REGION Network 18: I21.1 - Tank Group Pressure HIHI (PS-436)
   // True = OK, False = HIHI
   RUNG wire#powerrail
      I_Contact( "RIO2 Tanks Pressure Switch Hi Hi" )
      Coil( "20_TANKS_IP_DATA".RIO_02.FIRST_TANK.TANKS_PRESS_HIHI )
   END_RUNG
   // the same network as SCL:
   "20_TANKS_IP_DATA".RIO_02.FIRST_TANK.TANKS_PRESS_HIHI := NOT "RIO2 Tanks Pressure Switch Hi Hi";
END_REGION

REGION Network 19: I21.2 - Tank Level HIHI - (LS-425) - Second Tank
   // True = OK, False = HIHI
   RUNG wire#powerrail
      I_Contact( "Tank 2S BWT Level High High Switch" )
      Coil( "20_TANKS_IP_DATA".RIO_02.SECOND_TANK.BWT_LEVEL_HIHI )
   END_RUNG
   // the same network as SCL:
   "20_TANKS_IP_DATA".RIO_02.SECOND_TANK.BWT_LEVEL_HIHI := NOT "Tank 2S BWT Level High High Switch";
END_REGION

REGION Network 20: I21.3 - Spare Input
   // True = N/A, False = N/A
   RUNG wire#powerrail
      Contact( "RIO2_SPR_DI_21_3" )
      Coil( "20_TANKS_IP_DATA".RIO_02.FIRST_TANK.TANK_GROUP_SPARE_DI_3 )
   END_RUNG
   // the same network as SCL:
   "20_TANKS_IP_DATA".RIO_02.FIRST_TANK.TANK_GROUP_SPARE_DI_3 := "RIO2_SPR_DI_21_3";
END_REGION

REGION Network 21: I21.4 - Spare Input
   // True = N/A, False = N/A
   RUNG wire#powerrail
      Contact( "RIO2_SPR_DI_21_4" )
      Coil( "20_TANKS_IP_DATA".RIO_02.FIRST_TANK.TANK_GROUP_SPARE_DI_4 )
   END_RUNG
   // the same network as SCL:
   "20_TANKS_IP_DATA".RIO_02.FIRST_TANK.TANK_GROUP_SPARE_DI_4 := "RIO2_SPR_DI_21_4";
END_REGION

REGION Network 22: I21.5 - Spare Input
   // True = N/A, False = N/A
   RUNG wire#powerrail
      Contact( "RIO2_SPR_DI_21_5" )
      Coil( "20_TANKS_IP_DATA".RIO_02.FIRST_TANK.TANK_GROUP_SPARE_DI_5 )
   END_RUNG
   // the same network as SCL:
   "20_TANKS_IP_DATA".RIO_02.FIRST_TANK.TANK_GROUP_SPARE_DI_5 := "RIO2_SPR_DI_21_5";
END_REGION

REGION Network 23: I21.6 - Spare Input
   // True = N/A, False = N/A
   RUNG wire#powerrail
      Contact( "RIO2_SPR_DI_21_6" )
      Coil( "20_TANKS_IP_DATA".RIO_02.FIRST_TANK.TANK_GROUP_SPARE_DI_6 )
   END_RUNG
   // the same network as SCL:
   "20_TANKS_IP_DATA".RIO_02.FIRST_TANK.TANK_GROUP_SPARE_DI_6 := "RIO2_SPR_DI_21_6";
END_REGION

REGION Network 24: I21.7 - Spare Input
   // True = N/A, False = N/A
   RUNG wire#powerrail
      Contact( "RIO2_SPR_DI_21_7" )
      Coil( "20_TANKS_IP_DATA".RIO_02.FIRST_TANK.TANK_GROUP_SPARE_DI_7 )
   END_RUNG
   // the same network as SCL:
   "20_TANKS_IP_DATA".RIO_02.FIRST_TANK.TANK_GROUP_SPARE_DI_7 := "RIO2_SPR_DI_21_7";
END_REGION
END_FUNCTION

FUNCTION "23_RIO_3_DI_Processing" : Void   // FC23, LAD
TITLE = RIO Rack Digital Input Processing (Tank 1 = 3P, Tank 2 = 3S)
{ S7_Optimized_Access := 'TRUE' }
AUTHOR : JRS
VERSION : 0.1
// To process raw inputs prior to code use
BEGIN

REGION Network 1: I27.0 - Gas To Tank Valve Feedback Open (CV-422)
   // True = OPEN, False = NOT
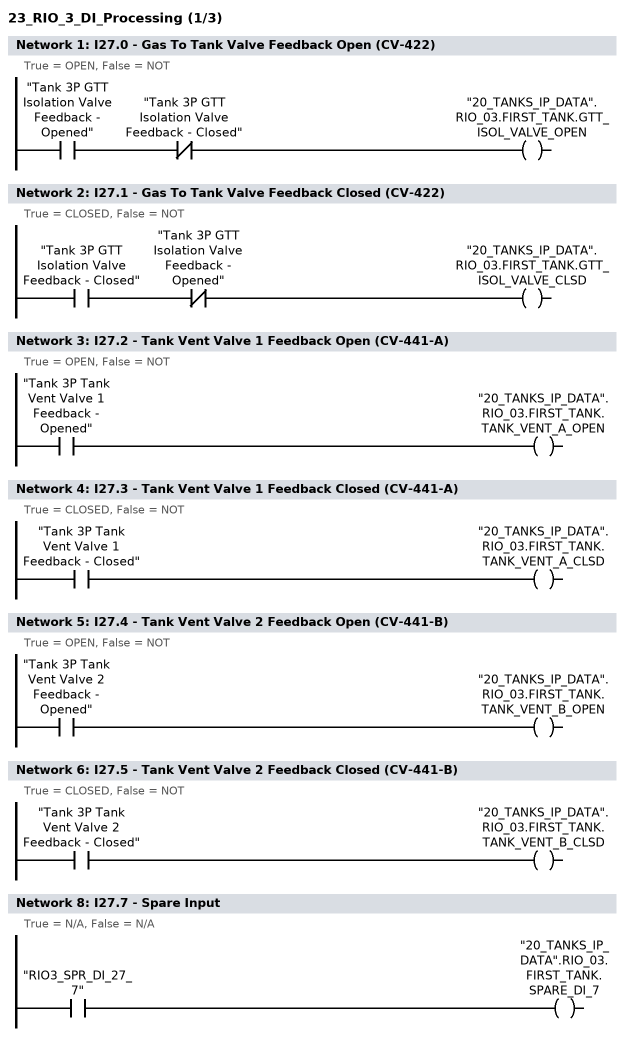
   RUNG wire#powerrail
      Contact( "Tank 3P GTT Isolation Valve Feedback - Opened" )
      I_Contact( "Tank 3P GTT Isolation Valve Feedback - Closed" )
      Coil( "20_TANKS_IP_DATA".RIO_03.FIRST_TANK.GTT_ISOL_VALVE_OPEN )
   END_RUNG
   // the same network as SCL:
   "20_TANKS_IP_DATA".RIO_03.FIRST_TANK.GTT_ISOL_VALVE_OPEN := "Tank 3P GTT Isolation Valve Feedback - Opened" AND NOT "Tank 3P GTT Isolation Valve Feedback - Closed";
END_REGION

REGION Network 2: I27.1 - Gas To Tank Valve Feedback Closed (CV-422)
   // True = CLOSED, False = NOT
   RUNG wire#powerrail
      Contact( "Tank 3P GTT Isolation Valve Feedback - Closed" )
      I_Contact( "Tank 3P GTT Isolation Valve Feedback - Opened" )
      Coil( "20_TANKS_IP_DATA".RIO_03.FIRST_TANK.GTT_ISOL_VALVE_CLSD )
   END_RUNG
   // the same network as SCL:
   "20_TANKS_IP_DATA".RIO_03.FIRST_TANK.GTT_ISOL_VALVE_CLSD := "Tank 3P GTT Isolation Valve Feedback - Closed" AND NOT "Tank 3P GTT Isolation Valve Feedback - Opened";
END_REGION

REGION Network 3: I27.2 - Tank Vent Valve 1 Feedback Open (CV-441-A)
   // True = OPEN, False = NOT
   RUNG wire#powerrail
      Contact( "Tank 3P Tank Vent Valve 1 Feedback - Opened" )
      Coil( "20_TANKS_IP_DATA".RIO_03.FIRST_TANK.TANK_VENT_A_OPEN )
   END_RUNG
   // the same network as SCL:
   "20_TANKS_IP_DATA".RIO_03.FIRST_TANK.TANK_VENT_A_OPEN := "Tank 3P Tank Vent Valve 1 Feedback - Opened";
END_REGION

REGION Network 4: I27.3 - Tank Vent Valve 1 Feedback Closed (CV-441-A)
   // True = CLOSED, False = NOT
   RUNG wire#powerrail
      Contact( "Tank 3P Tank Vent Valve 1 Feedback - Closed" )
      Coil( "20_TANKS_IP_DATA".RIO_03.FIRST_TANK.TANK_VENT_A_CLSD )
   END_RUNG
   // the same network as SCL:
   "20_TANKS_IP_DATA".RIO_03.FIRST_TANK.TANK_VENT_A_CLSD := "Tank 3P Tank Vent Valve 1 Feedback - Closed";
END_REGION

REGION Network 5: I27.4 - Tank Vent Valve 2 Feedback Open (CV-441-B)
   // True = OPEN, False = NOT
   RUNG wire#powerrail
      Contact( "Tank 3P Tank Vent Valve 2 Feedback - Opened" )
      Coil( "20_TANKS_IP_DATA".RIO_03.FIRST_TANK.TANK_VENT_B_OPEN )
   END_RUNG
   // the same network as SCL:
   "20_TANKS_IP_DATA".RIO_03.FIRST_TANK.TANK_VENT_B_OPEN := "Tank 3P Tank Vent Valve 2 Feedback - Opened";
END_REGION

REGION Network 6: I27.5 - Tank Vent Valve 2 Feedback Closed (CV-441-B)
   // True = CLOSED, False = NOT
   RUNG wire#powerrail
      Contact( "Tank 3P Tank Vent Valve 2 Feedback - Closed" )
      Coil( "20_TANKS_IP_DATA".RIO_03.FIRST_TANK.TANK_VENT_B_CLSD )
   END_RUNG
   // the same network as SCL:
   "20_TANKS_IP_DATA".RIO_03.FIRST_TANK.TANK_VENT_B_CLSD := "Tank 3P Tank Vent Valve 2 Feedback - Closed";
END_REGION

REGION Network 7: I27.6 - Spare Input Accesed from Warning FC
   // True = N/A, False = N/A
END_REGION

REGION Network 8: I27.7 - Spare Input
   // True = N/A, False = N/A
   RUNG wire#powerrail
      Contact( "RIO3_SPR_DI_27_7" )
      Coil( "20_TANKS_IP_DATA".RIO_03.FIRST_TANK.SPARE_DI_7 )
   END_RUNG
   // the same network as SCL:
   "20_TANKS_IP_DATA".RIO_03.FIRST_TANK.SPARE_DI_7 := "RIO3_SPR_DI_27_7";
END_REGION

REGION Network 9: I30.0 - Gas To Tank Valve Feedback Open (CV-422)
   // True = OPEN, False = NOT
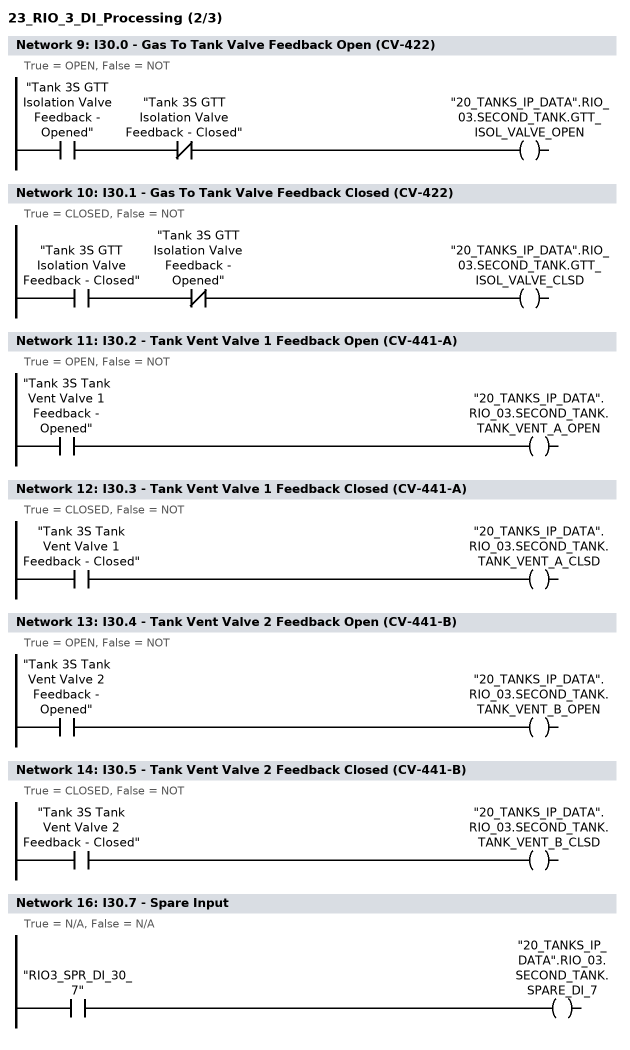
   RUNG wire#powerrail
      Contact( "Tank 3S GTT Isolation Valve Feedback - Opened" )
      I_Contact( "Tank 3S GTT Isolation Valve Feedback - Closed" )
      Coil( "20_TANKS_IP_DATA".RIO_03.SECOND_TANK.GTT_ISOL_VALVE_OPEN )
   END_RUNG
   // the same network as SCL:
   "20_TANKS_IP_DATA".RIO_03.SECOND_TANK.GTT_ISOL_VALVE_OPEN := "Tank 3S GTT Isolation Valve Feedback - Opened" AND NOT "Tank 3S GTT Isolation Valve Feedback - Closed";
END_REGION

REGION Network 10: I30.1 - Gas To Tank Valve Feedback Closed (CV-422)
   // True = CLOSED, False = NOT
   RUNG wire#powerrail
      Contact( "Tank 3S GTT Isolation Valve Feedback - Closed" )
      I_Contact( "Tank 3S GTT Isolation Valve Feedback - Opened" )
      Coil( "20_TANKS_IP_DATA".RIO_03.SECOND_TANK.GTT_ISOL_VALVE_CLSD )
   END_RUNG
   // the same network as SCL:
   "20_TANKS_IP_DATA".RIO_03.SECOND_TANK.GTT_ISOL_VALVE_CLSD := "Tank 3S GTT Isolation Valve Feedback - Closed" AND NOT "Tank 3S GTT Isolation Valve Feedback - Opened";
END_REGION

REGION Network 11: I30.2 - Tank Vent Valve 1 Feedback Open (CV-441-A)
   // True = OPEN, False = NOT
   RUNG wire#powerrail
      Contact( "Tank 3S Tank Vent Valve 1 Feedback - Opened" )
      Coil( "20_TANKS_IP_DATA".RIO_03.SECOND_TANK.TANK_VENT_A_OPEN )
   END_RUNG
   // the same network as SCL:
   "20_TANKS_IP_DATA".RIO_03.SECOND_TANK.TANK_VENT_A_OPEN := "Tank 3S Tank Vent Valve 1 Feedback - Opened";
END_REGION

REGION Network 12: I30.3 - Tank Vent Valve 1 Feedback Closed (CV-441-A)
   // True = CLOSED, False = NOT
   RUNG wire#powerrail
      Contact( "Tank 3S Tank Vent Valve 1 Feedback - Closed" )
      Coil( "20_TANKS_IP_DATA".RIO_03.SECOND_TANK.TANK_VENT_A_CLSD )
   END_RUNG
   // the same network as SCL:
   "20_TANKS_IP_DATA".RIO_03.SECOND_TANK.TANK_VENT_A_CLSD := "Tank 3S Tank Vent Valve 1 Feedback - Closed";
END_REGION

REGION Network 13: I30.4 - Tank Vent Valve 2 Feedback Open (CV-441-B)
   // True = OPEN, False = NOT
   RUNG wire#powerrail
      Contact( "Tank 3S Tank Vent Valve 2 Feedback - Opened" )
      Coil( "20_TANKS_IP_DATA".RIO_03.SECOND_TANK.TANK_VENT_B_OPEN )
   END_RUNG
   // the same network as SCL:
   "20_TANKS_IP_DATA".RIO_03.SECOND_TANK.TANK_VENT_B_OPEN := "Tank 3S Tank Vent Valve 2 Feedback - Opened";
END_REGION

REGION Network 14: I30.5 - Tank Vent Valve 2 Feedback Closed (CV-441-B)
   // True = CLOSED, False = NOT
   RUNG wire#powerrail
      Contact( "Tank 3S Tank Vent Valve 2 Feedback - Closed" )
      Coil( "20_TANKS_IP_DATA".RIO_03.SECOND_TANK.TANK_VENT_B_CLSD )
   END_RUNG
   // the same network as SCL:
   "20_TANKS_IP_DATA".RIO_03.SECOND_TANK.TANK_VENT_B_CLSD := "Tank 3S Tank Vent Valve 2 Feedback - Closed";
END_REGION

REGION Network 15: I30.6 - Spare Input Accesed from Warning FC
   // True = N/A, False = N/A
END_REGION

REGION Network 16: I30.7 - Spare Input
   // True = N/A, False = N/A
   RUNG wire#powerrail
      Contact( "RIO3_SPR_DI_30_7" )
      Coil( "20_TANKS_IP_DATA".RIO_03.SECOND_TANK.SPARE_DI_7 )
   END_RUNG
   // the same network as SCL:
   "20_TANKS_IP_DATA".RIO_03.SECOND_TANK.SPARE_DI_7 := "RIO3_SPR_DI_30_7";
END_REGION

REGION Network 17: I33.0 - Tank Level HIHI - (LS-425) - First Tank
   // True = OK, False = HIHI
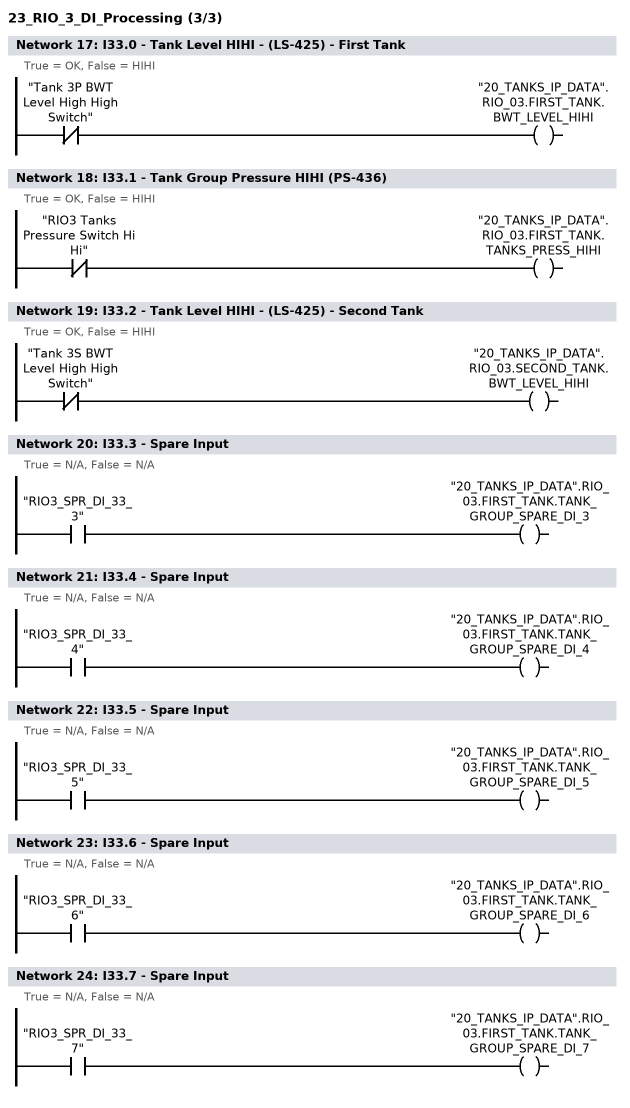
   RUNG wire#powerrail
      I_Contact( "Tank 3P BWT Level High High Switch" )
      Coil( "20_TANKS_IP_DATA".RIO_03.FIRST_TANK.BWT_LEVEL_HIHI )
   END_RUNG
   // the same network as SCL:
   "20_TANKS_IP_DATA".RIO_03.FIRST_TANK.BWT_LEVEL_HIHI := NOT "Tank 3P BWT Level High High Switch";
END_REGION

REGION Network 18: I33.1 - Tank Group Pressure HIHI (PS-436)
   // True = OK, False = HIHI
   RUNG wire#powerrail
      I_Contact( "RIO3 Tanks Pressure Switch Hi Hi" )
      Coil( "20_TANKS_IP_DATA".RIO_03.FIRST_TANK.TANKS_PRESS_HIHI )
   END_RUNG
   // the same network as SCL:
   "20_TANKS_IP_DATA".RIO_03.FIRST_TANK.TANKS_PRESS_HIHI := NOT "RIO3 Tanks Pressure Switch Hi Hi";
END_REGION

REGION Network 19: I33.2 - Tank Level HIHI - (LS-425) - Second Tank
   // True = OK, False = HIHI
   RUNG wire#powerrail
      I_Contact( "Tank 3S BWT Level High High Switch" )
      Coil( "20_TANKS_IP_DATA".RIO_03.SECOND_TANK.BWT_LEVEL_HIHI )
   END_RUNG
   // the same network as SCL:
   "20_TANKS_IP_DATA".RIO_03.SECOND_TANK.BWT_LEVEL_HIHI := NOT "Tank 3S BWT Level High High Switch";
END_REGION

REGION Network 20: I33.3 - Spare Input
   // True = N/A, False = N/A
   RUNG wire#powerrail
      Contact( "RIO3_SPR_DI_33_3" )
      Coil( "20_TANKS_IP_DATA".RIO_03.FIRST_TANK.TANK_GROUP_SPARE_DI_3 )
   END_RUNG
   // the same network as SCL:
   "20_TANKS_IP_DATA".RIO_03.FIRST_TANK.TANK_GROUP_SPARE_DI_3 := "RIO3_SPR_DI_33_3";
END_REGION

REGION Network 21: I33.4 - Spare Input
   // True = N/A, False = N/A
   RUNG wire#powerrail
      Contact( "RIO3_SPR_DI_33_4" )
      Coil( "20_TANKS_IP_DATA".RIO_03.FIRST_TANK.TANK_GROUP_SPARE_DI_4 )
   END_RUNG
   // the same network as SCL:
   "20_TANKS_IP_DATA".RIO_03.FIRST_TANK.TANK_GROUP_SPARE_DI_4 := "RIO3_SPR_DI_33_4";
END_REGION

REGION Network 22: I33.5 - Spare Input
   // True = N/A, False = N/A
   RUNG wire#powerrail
      Contact( "RIO3_SPR_DI_33_5" )
      Coil( "20_TANKS_IP_DATA".RIO_03.FIRST_TANK.TANK_GROUP_SPARE_DI_5 )
   END_RUNG
   // the same network as SCL:
   "20_TANKS_IP_DATA".RIO_03.FIRST_TANK.TANK_GROUP_SPARE_DI_5 := "RIO3_SPR_DI_33_5";
END_REGION

REGION Network 23: I33.6 - Spare Input
   // True = N/A, False = N/A
   RUNG wire#powerrail
      Contact( "RIO3_SPR_DI_33_6" )
      Coil( "20_TANKS_IP_DATA".RIO_03.FIRST_TANK.TANK_GROUP_SPARE_DI_6 )
   END_RUNG
   // the same network as SCL:
   "20_TANKS_IP_DATA".RIO_03.FIRST_TANK.TANK_GROUP_SPARE_DI_6 := "RIO3_SPR_DI_33_6";
END_REGION

REGION Network 24: I33.7 - Spare Input
   // True = N/A, False = N/A
   RUNG wire#powerrail
      Contact( "RIO3_SPR_DI_33_7" )
      Coil( "20_TANKS_IP_DATA".RIO_03.FIRST_TANK.TANK_GROUP_SPARE_DI_7 )
   END_RUNG
   // the same network as SCL:
   "20_TANKS_IP_DATA".RIO_03.FIRST_TANK.TANK_GROUP_SPARE_DI_7 := "RIO3_SPR_DI_33_7";
END_REGION
END_FUNCTION

FUNCTION "24_RIO_4_DI_Processing" : Void   // FC24, LAD
TITLE = RIO Rack Digital Input Processing (Tank 1 = 4P, Tank 2 = 4S)
{ S7_Optimized_Access := 'TRUE' }
AUTHOR : JRS
VERSION : 0.1
// To process raw inputs prior to code use
BEGIN

REGION Network 1: I39.0 - Gas To Tank Valve Feedback Open (CV-422)
   // True = OPEN, False = NOT
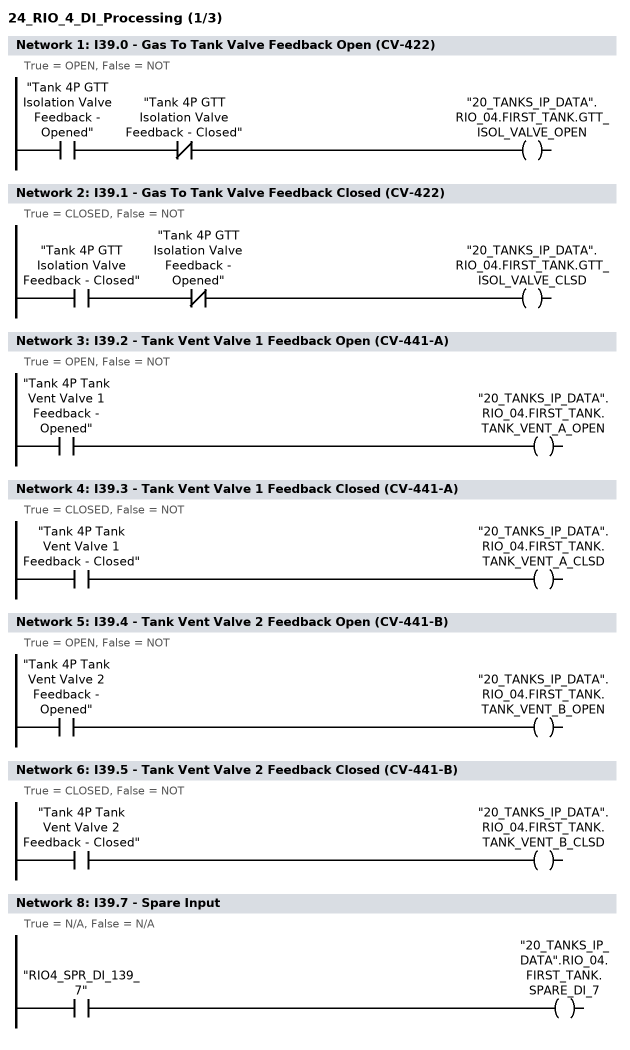
   RUNG wire#powerrail
      Contact( "Tank 4P GTT Isolation Valve Feedback - Opened" )
      I_Contact( "Tank 4P GTT Isolation Valve Feedback - Closed" )
      Coil( "20_TANKS_IP_DATA".RIO_04.FIRST_TANK.GTT_ISOL_VALVE_OPEN )
   END_RUNG
   // the same network as SCL:
   "20_TANKS_IP_DATA".RIO_04.FIRST_TANK.GTT_ISOL_VALVE_OPEN := "Tank 4P GTT Isolation Valve Feedback - Opened" AND NOT "Tank 4P GTT Isolation Valve Feedback - Closed";
END_REGION

REGION Network 2: I39.1 - Gas To Tank Valve Feedback Closed (CV-422)
   // True = CLOSED, False = NOT
   RUNG wire#powerrail
      Contact( "Tank 4P GTT Isolation Valve Feedback - Closed" )
      I_Contact( "Tank 4P GTT Isolation Valve Feedback - Opened" )
      Coil( "20_TANKS_IP_DATA".RIO_04.FIRST_TANK.GTT_ISOL_VALVE_CLSD )
   END_RUNG
   // the same network as SCL:
   "20_TANKS_IP_DATA".RIO_04.FIRST_TANK.GTT_ISOL_VALVE_CLSD := "Tank 4P GTT Isolation Valve Feedback - Closed" AND NOT "Tank 4P GTT Isolation Valve Feedback - Opened";
END_REGION

REGION Network 3: I39.2 - Tank Vent Valve 1 Feedback Open (CV-441-A)
   // True = OPEN, False = NOT
   RUNG wire#powerrail
      Contact( "Tank 4P Tank Vent Valve 1 Feedback - Opened" )
      Coil( "20_TANKS_IP_DATA".RIO_04.FIRST_TANK.TANK_VENT_A_OPEN )
   END_RUNG
   // the same network as SCL:
   "20_TANKS_IP_DATA".RIO_04.FIRST_TANK.TANK_VENT_A_OPEN := "Tank 4P Tank Vent Valve 1 Feedback - Opened";
END_REGION

REGION Network 4: I39.3 - Tank Vent Valve 1 Feedback Closed (CV-441-A)
   // True = CLOSED, False = NOT
   RUNG wire#powerrail
      Contact( "Tank 4P Tank Vent Valve 1 Feedback - Closed" )
      Coil( "20_TANKS_IP_DATA".RIO_04.FIRST_TANK.TANK_VENT_A_CLSD )
   END_RUNG
   // the same network as SCL:
   "20_TANKS_IP_DATA".RIO_04.FIRST_TANK.TANK_VENT_A_CLSD := "Tank 4P Tank Vent Valve 1 Feedback - Closed";
END_REGION

REGION Network 5: I39.4 - Tank Vent Valve 2 Feedback Open (CV-441-B)
   // True = OPEN, False = NOT
   RUNG wire#powerrail
      Contact( "Tank 4P Tank Vent Valve 2 Feedback - Opened" )
      Coil( "20_TANKS_IP_DATA".RIO_04.FIRST_TANK.TANK_VENT_B_OPEN )
   END_RUNG
   // the same network as SCL:
   "20_TANKS_IP_DATA".RIO_04.FIRST_TANK.TANK_VENT_B_OPEN := "Tank 4P Tank Vent Valve 2 Feedback - Opened";
END_REGION

REGION Network 6: I39.5 - Tank Vent Valve 2 Feedback Closed (CV-441-B)
   // True = CLOSED, False = NOT
   RUNG wire#powerrail
      Contact( "Tank 4P Tank Vent Valve 2 Feedback - Closed" )
      Coil( "20_TANKS_IP_DATA".RIO_04.FIRST_TANK.TANK_VENT_B_CLSD )
   END_RUNG
   // the same network as SCL:
   "20_TANKS_IP_DATA".RIO_04.FIRST_TANK.TANK_VENT_B_CLSD := "Tank 4P Tank Vent Valve 2 Feedback - Closed";
END_REGION

REGION Network 7: I39.6 - Spare Input Destination Accesed from Warning FC
   // True = N/A, False = N/A
END_REGION

REGION Network 8: I39.7 - Spare Input
   // True = N/A, False = N/A
   RUNG wire#powerrail
      Contact( "RIO4_SPR_DI_139_7" )
      Coil( "20_TANKS_IP_DATA".RIO_04.FIRST_TANK.SPARE_DI_7 )
   END_RUNG
   // the same network as SCL:
   "20_TANKS_IP_DATA".RIO_04.FIRST_TANK.SPARE_DI_7 := "RIO4_SPR_DI_139_7";
END_REGION

REGION Network 9: I42.0 - Gas To Tank Valve Feedback Open (CV-422)
   // True = OPEN, False = NOT
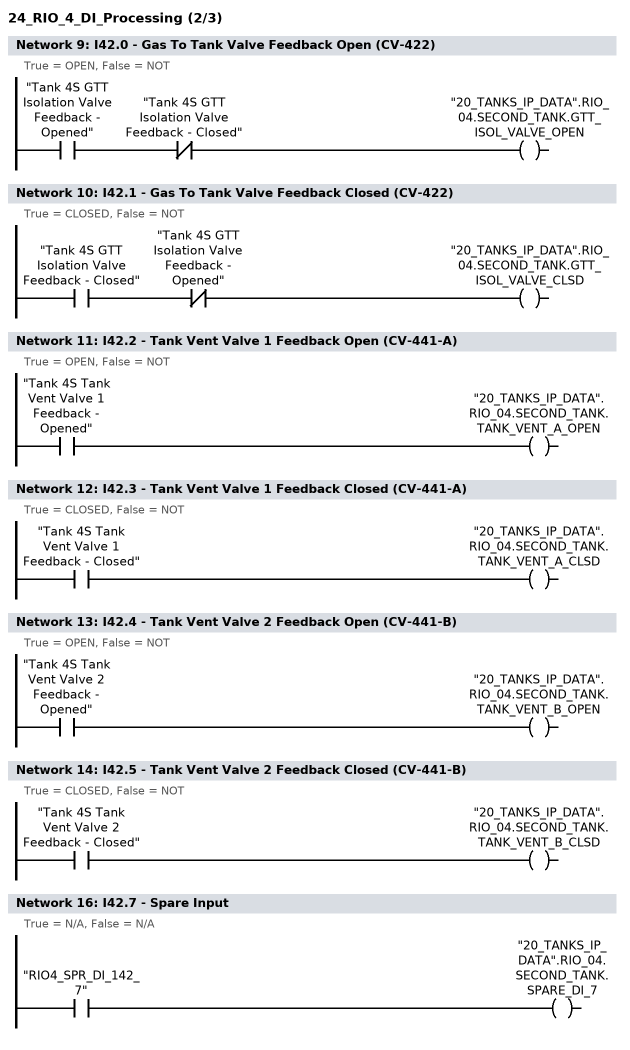
   RUNG wire#powerrail
      Contact( "Tank 4S GTT Isolation Valve Feedback - Opened" )
      I_Contact( "Tank 4S GTT Isolation Valve Feedback - Closed" )
      Coil( "20_TANKS_IP_DATA".RIO_04.SECOND_TANK.GTT_ISOL_VALVE_OPEN )
   END_RUNG
   // the same network as SCL:
   "20_TANKS_IP_DATA".RIO_04.SECOND_TANK.GTT_ISOL_VALVE_OPEN := "Tank 4S GTT Isolation Valve Feedback - Opened" AND NOT "Tank 4S GTT Isolation Valve Feedback - Closed";
END_REGION

REGION Network 10: I42.1 - Gas To Tank Valve Feedback Closed (CV-422)
   // True = CLOSED, False = NOT
   RUNG wire#powerrail
      Contact( "Tank 4S GTT Isolation Valve Feedback - Closed" )
      I_Contact( "Tank 4S GTT Isolation Valve Feedback - Opened" )
      Coil( "20_TANKS_IP_DATA".RIO_04.SECOND_TANK.GTT_ISOL_VALVE_CLSD )
   END_RUNG
   // the same network as SCL:
   "20_TANKS_IP_DATA".RIO_04.SECOND_TANK.GTT_ISOL_VALVE_CLSD := "Tank 4S GTT Isolation Valve Feedback - Closed" AND NOT "Tank 4S GTT Isolation Valve Feedback - Opened";
END_REGION

REGION Network 11: I42.2 - Tank Vent Valve 1 Feedback Open (CV-441-A)
   // True = OPEN, False = NOT
   RUNG wire#powerrail
      Contact( "Tank 4S Tank Vent Valve 1 Feedback - Opened" )
      Coil( "20_TANKS_IP_DATA".RIO_04.SECOND_TANK.TANK_VENT_A_OPEN )
   END_RUNG
   // the same network as SCL:
   "20_TANKS_IP_DATA".RIO_04.SECOND_TANK.TANK_VENT_A_OPEN := "Tank 4S Tank Vent Valve 1 Feedback - Opened";
END_REGION

REGION Network 12: I42.3 - Tank Vent Valve 1 Feedback Closed (CV-441-A)
   // True = CLOSED, False = NOT
   RUNG wire#powerrail
      Contact( "Tank 4S Tank Vent Valve 1 Feedback - Closed" )
      Coil( "20_TANKS_IP_DATA".RIO_04.SECOND_TANK.TANK_VENT_A_CLSD )
   END_RUNG
   // the same network as SCL:
   "20_TANKS_IP_DATA".RIO_04.SECOND_TANK.TANK_VENT_A_CLSD := "Tank 4S Tank Vent Valve 1 Feedback - Closed";
END_REGION

REGION Network 13: I42.4 - Tank Vent Valve 2 Feedback Open (CV-441-B)
   // True = OPEN, False = NOT
   RUNG wire#powerrail
      Contact( "Tank 4S Tank Vent Valve 2 Feedback - Opened" )
      Coil( "20_TANKS_IP_DATA".RIO_04.SECOND_TANK.TANK_VENT_B_OPEN )
   END_RUNG
   // the same network as SCL:
   "20_TANKS_IP_DATA".RIO_04.SECOND_TANK.TANK_VENT_B_OPEN := "Tank 4S Tank Vent Valve 2 Feedback - Opened";
END_REGION

